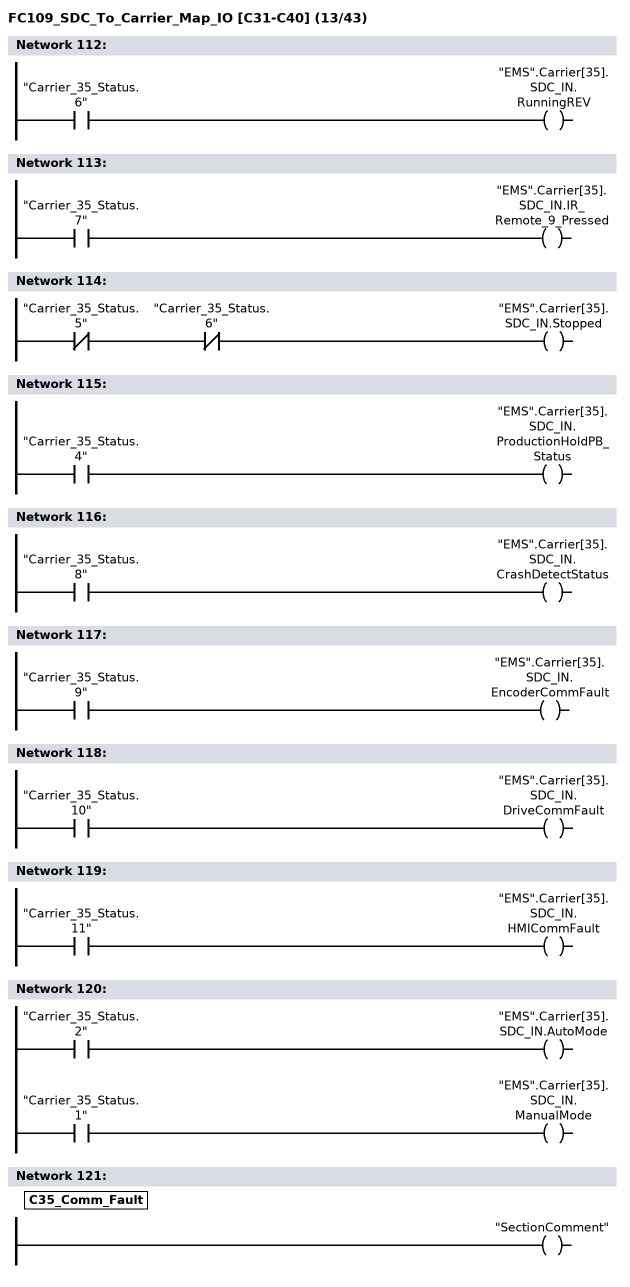
   RUNG wire#powerrail
      Contact( "Carrier_35_Status.6" )
      Coil( "EMS".Carrier[35].SDC_IN.RunningREV )
   END_RUNG
   // the same network as SCL:
   "EMS".Carrier[35].SDC_IN.RunningREV := "Carrier_35_Status.6";
END_REGION

REGION Network 113
   RUNG wire#powerrail
      Contact( "Carrier_35_Status.7" )
      Coil( "EMS".Carrier[35].SDC_IN.IR_Remote_9_Pressed )
   END_RUNG
   // the same network as SCL:
   "EMS".Carrier[35].SDC_IN.IR_Remote_9_Pressed := "Carrier_35_Status.7";
END_REGION

REGION Network 114
   RUNG wire#powerrail
      I_Contact( "Carrier_35_Status.5" )
      I_Contact( "Carrier_35_Status.6" )
      Coil( "EMS".Carrier[35].SDC_IN.Stopped )
   END_RUNG
   // the same network as SCL:
   "EMS".Carrier[35].SDC_IN.Stopped := NOT "Carrier_35_Status.5" AND NOT "Carrier_35_Status.6";
END_REGION

REGION Network 115
   RUNG wire#powerrail
      Contact( "Carrier_35_Status.4" )
      Coil( "EMS".Carrier[35].SDC_IN.ProductionHoldPB_Status )
   END_RUNG
   // the same network as SCL:
   "EMS".Carrier[35].SDC_IN.ProductionHoldPB_Status := "Carrier_35_Status.4";
END_REGION

REGION Network 116
   RUNG wire#powerrail
      Contact( "Carrier_35_Status.8" )
      Coil( "EMS".Carrier[35].SDC_IN.CrashDetectStatus )
   END_RUNG
   // the same network as SCL:
   "EMS".Carrier[35].SDC_IN.CrashDetectStatus := "Carrier_35_Status.8";
END_REGION

REGION Network 117
   RUNG wire#powerrail
      Contact( "Carrier_35_Status.9" )
      Coil( "EMS".Carrier[35].SDC_IN.EncoderCommFault )
   END_RUNG
   // the same network as SCL:
   "EMS".Carrier[35].SDC_IN.EncoderCommFault := "Carrier_35_Status.9";
END_REGION

REGION Network 118
   RUNG wire#powerrail
      Contact( "Carrier_35_Status.10" )
      Coil( "EMS".Carrier[35].SDC_IN.DriveCommFault )
   END_RUNG
   // the same network as SCL:
   "EMS".Carrier[35].SDC_IN.DriveCommFault := "Carrier_35_Status.10";
END_REGION

REGION Network 119
   RUNG wire#powerrail
      Contact( "Carrier_35_Status.11" )
      Coil( "EMS".Carrier[35].SDC_IN.HMICommFault )
   END_RUNG
   // the same network as SCL:
   "EMS".Carrier[35].SDC_IN.HMICommFault := "Carrier_35_Status.11";
END_REGION

REGION Network 120
   RUNG wire#powerrail
      Contact( "Carrier_35_Status.2" )
      Coil( "EMS".Carrier[35].SDC_IN.AutoMode )
   END_RUNG
   RUNG wire#powerrail
      Contact( "Carrier_35_Status.1" )
      Coil( "EMS".Carrier[35].SDC_IN.ManualMode )
   END_RUNG
   // the same network as SCL:
   "EMS".Carrier[35].SDC_IN.AutoMode := "Carrier_35_Status.2";
   "EMS".Carrier[35].SDC_IN.ManualMode := "Carrier_35_Status.1";
END_REGION

REGION Network 121
   Label( C35_Comm_Fault )
   RUNG wire#powerrail
      Coil( "SectionComment" )
   END_RUNG
   // the same network as SCL:
   C35_Comm_Fault:
   "SectionComment" := TRUE;
END_REGION

REGION Network 122
   // **********************************************************************************************************************
   // 
   // Carrier 36 I-Device Data Transfer Interlocks from Carrier to SDC
   // 
   // **********************************************************************************************************************
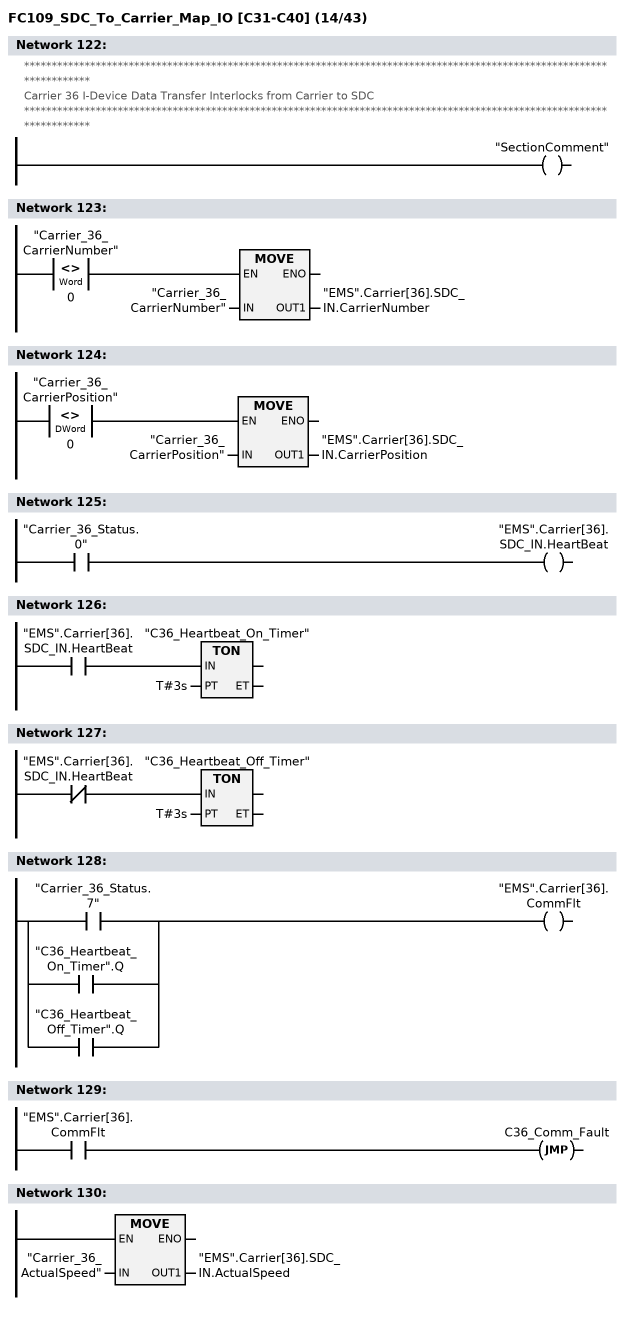
   RUNG wire#powerrail
      Coil( "SectionComment" )
   END_RUNG
   // the same network as SCL:
   "SectionComment" := TRUE;
END_REGION

REGION Network 123
   RUNG wire#powerrail
      { S7_Templates := "SrcType := Word" } NE_Contact(in1 := "Carrier_36_CarrierNumber", in2 := 0)
      Move(in := "Carrier_36_CarrierNumber", out1 => "EMS".Carrier[36].SDC_IN.CarrierNumber)
   END_RUNG
   // the same network as SCL:
   IF "Carrier_36_CarrierNumber" <> 0 THEN
       "EMS".Carrier[36].SDC_IN.CarrierNumber := "Carrier_36_CarrierNumber";
   END_IF;
END_REGION

REGION Network 124
   RUNG wire#powerrail
      { S7_Templates := "SrcType := DWord" } NE_Contact(in1 := "Carrier_36_CarrierPosition", in2 := 0)
      Move(in := "Carrier_36_CarrierPosition", out1 => "EMS".Carrier[36].SDC_IN.CarrierPosition)
   END_RUNG
   // the same network as SCL:
   IF "Carrier_36_CarrierPosition" <> 0 THEN
       "EMS".Carrier[36].SDC_IN.CarrierPosition := "Carrier_36_CarrierPosition";
   END_IF;
END_REGION

REGION Network 125
   RUNG wire#powerrail
      Contact( "Carrier_36_Status.0" )
      Coil( "EMS".Carrier[36].SDC_IN.HeartBeat )
   END_RUNG
   // the same network as SCL:
   "EMS".Carrier[36].SDC_IN.HeartBeat := "Carrier_36_Status.0";
END_REGION

REGION Network 126
   "C36_Heartbeat_On_Timer".TON(IN := "EMS".Carrier[36].SDC_IN.HeartBeat, PT := T#3s);
END_REGION

REGION Network 127
   "C36_Heartbeat_Off_Timer".TON(IN := NOT "EMS".Carrier[36].SDC_IN.HeartBeat, PT := T#3s);
END_REGION

REGION Network 128
   RUNG wire#powerrail
      Contact( "Carrier_36_Status.7" )
      wire#w1
      Coil( "EMS".Carrier[36].CommFlt )
   END_RUNG
   RUNG wire#powerrail
      Contact( "C36_Heartbeat_On_Timer".Q )
   END_RUNG wire#w1
   RUNG wire#powerrail
      Contact( "C36_Heartbeat_Off_Timer".Q )
   END_RUNG wire#w1
   // the same network as SCL:
   "EMS".Carrier[36].CommFlt := "Carrier_36_Status.7" OR "C36_Heartbeat_On_Timer".Q OR "C36_Heartbeat_Off_Timer".Q;
END_REGION

REGION Network 129
   RUNG wire#powerrail
      Contact( "EMS".Carrier[36].CommFlt )
      JumpCoil( C36_Comm_Fault )
   END_RUNG
   // the same network as SCL:
   IF "EMS".Carrier[36].CommFlt THEN GOTO C36_Comm_Fault; END_IF;
END_REGION

REGION Network 130
   RUNG wire#powerrail
      Move(in := "Carrier_36_ActualSpeed", out1 => "EMS".Carrier[36].SDC_IN.ActualSpeed)
   END_RUNG
   // the same network as SCL:
   "EMS".Carrier[36].SDC_IN.ActualSpeed := "Carrier_36_ActualSpeed";
END_REGION

REGION Network 131
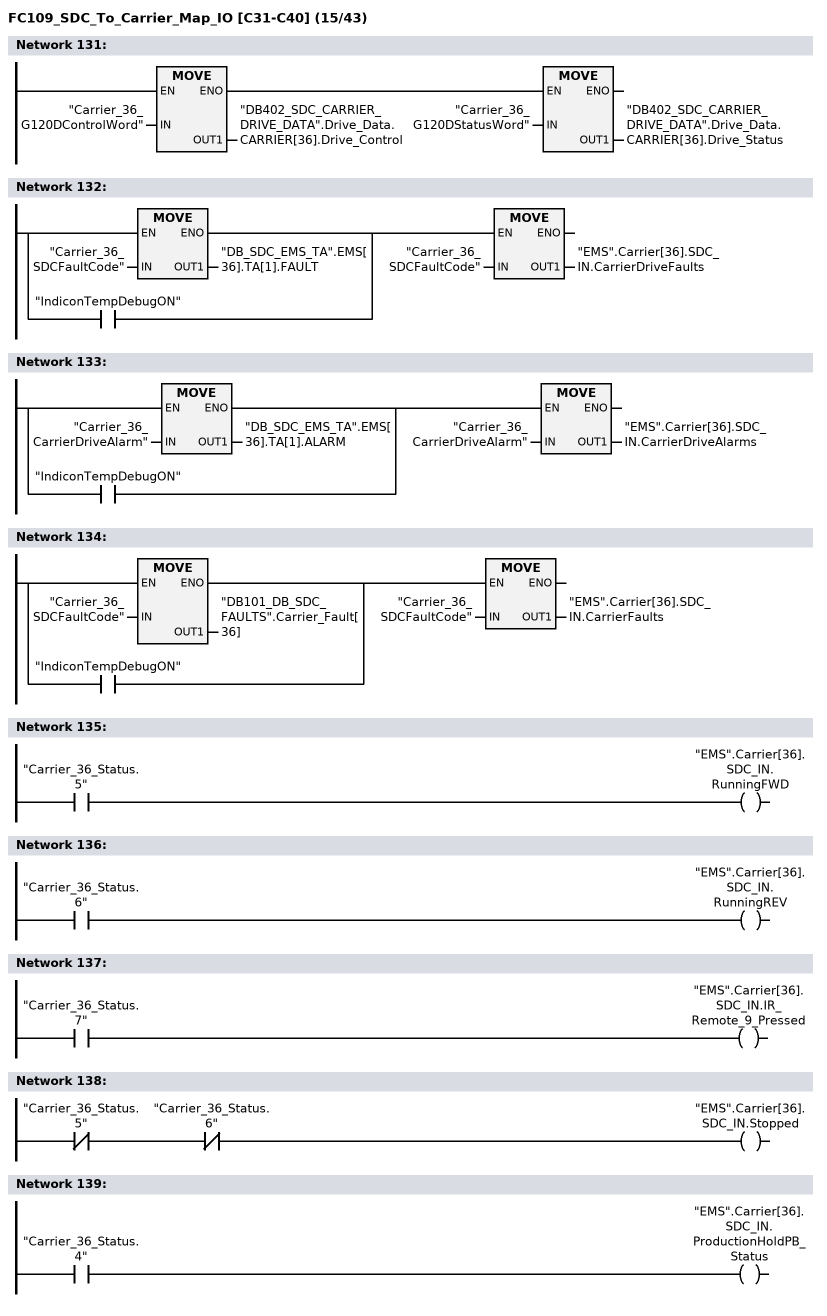
   RUNG wire#powerrail
      Move(in := "Carrier_36_G120DControlWord", out1 => "DB402_SDC_CARRIER_DRIVE_DATA".Drive_Data.CARRIER[36].Drive_Control)
      Move(in := "Carrier_36_G120DStatusWord", out1 => "DB402_SDC_CARRIER_DRIVE_DATA".Drive_Data.CARRIER[36].Drive_Status)
   END_RUNG
   // the same network as SCL:
   "DB402_SDC_CARRIER_DRIVE_DATA".Drive_Data.CARRIER[36].Drive_Control := "Carrier_36_G120DControlWord";
   "DB402_SDC_CARRIER_DRIVE_DATA".Drive_Data.CARRIER[36].Drive_Status := "Carrier_36_G120DStatusWord";
END_REGION

REGION Network 132
   RUNG wire#powerrail
      Move(in := "Carrier_36_SDCFaultCode", out1 => "DB_SDC_EMS_TA".EMS[36].TA[1].FAULT)
      wire#w1
      Move(in := "Carrier_36_SDCFaultCode", out1 => "EMS".Carrier[36].SDC_IN.CarrierDriveFaults)
   END_RUNG
   RUNG wire#powerrail
      Contact( "IndiconTempDebugON" )
   END_RUNG wire#w1
   // the same network as SCL:
   "DB_SDC_EMS_TA".EMS[36].TA[1].FAULT := "Carrier_36_SDCFaultCode";
   IF TRUE OR "IndiconTempDebugON" THEN
       "EMS".Carrier[36].SDC_IN.CarrierDriveFaults := "Carrier_36_SDCFaultCode";
   END_IF;
END_REGION

REGION Network 133
   RUNG wire#powerrail
      Move(in := "Carrier_36_CarrierDriveAlarm", out1 => "DB_SDC_EMS_TA".EMS[36].TA[1].ALARM)
      wire#w1
      Move(in := "Carrier_36_CarrierDriveAlarm", out1 => "EMS".Carrier[36].SDC_IN.CarrierDriveAlarms)
   END_RUNG
   RUNG wire#powerrail
      Contact( "IndiconTempDebugON" )
   END_RUNG wire#w1
   // the same network as SCL:
   "DB_SDC_EMS_TA".EMS[36].TA[1].ALARM := "Carrier_36_CarrierDriveAlarm";
   IF TRUE OR "IndiconTempDebugON" THEN
       "EMS".Carrier[36].SDC_IN.CarrierDriveAlarms := "Carrier_36_CarrierDriveAlarm";
   END_IF;
END_REGION

REGION Network 134
   RUNG wire#powerrail
      Move(in := "Carrier_36_SDCFaultCode", out1 => "DB101_DB_SDC_FAULTS".Carrier_Fault[36])
      wire#w1
      Move(in := "Carrier_36_SDCFaultCode", out1 => "EMS".Carrier[36].SDC_IN.CarrierFaults)
   END_RUNG
   RUNG wire#powerrail
      Contact( "IndiconTempDebugON" )
   END_RUNG wire#w1
   // the same network as SCL:
   "DB101_DB_SDC_FAULTS".Carrier_Fault[36] := "Carrier_36_SDCFaultCode";
   IF TRUE OR "IndiconTempDebugON" THEN
       "EMS".Carrier[36].SDC_IN.CarrierFaults := "Carrier_36_SDCFaultCode";
   END_IF;
END_REGION

REGION Network 135
   RUNG wire#powerrail
      Contact( "Carrier_36_Status.5" )
      Coil( "EMS".Carrier[36].SDC_IN.RunningFWD )
   END_RUNG
   // the same network as SCL:
   "EMS".Carrier[36].SDC_IN.RunningFWD := "Carrier_36_Status.5";
END_REGION

REGION Network 136
   RUNG wire#powerrail
      Contact( "Carrier_36_Status.6" )
      Coil( "EMS".Carrier[36].SDC_IN.RunningREV )
   END_RUNG
   // the same network as SCL:
   "EMS".Carrier[36].SDC_IN.RunningREV := "Carrier_36_Status.6";
END_REGION

REGION Network 137
   RUNG wire#powerrail
      Contact( "Carrier_36_Status.7" )
      Coil( "EMS".Carrier[36].SDC_IN.IR_Remote_9_Pressed )
   END_RUNG
   // the same network as SCL:
   "EMS".Carrier[36].SDC_IN.IR_Remote_9_Pressed := "Carrier_36_Status.7";
END_REGION

REGION Network 138
   RUNG wire#powerrail
      I_Contact( "Carrier_36_Status.5" )
      I_Contact( "Carrier_36_Status.6" )
      Coil( "EMS".Carrier[36].SDC_IN.Stopped )
   END_RUNG
   // the same network as SCL:
   "EMS".Carrier[36].SDC_IN.Stopped := NOT "Carrier_36_Status.5" AND NOT "Carrier_36_Status.6";
END_REGION

REGION Network 139
   RUNG wire#powerrail
      Contact( "Carrier_36_Status.4" )
      Coil( "EMS".Carrier[36].SDC_IN.ProductionHoldPB_Status )
   END_RUNG
   // the same network as SCL:
   "EMS".Carrier[36].SDC_IN.ProductionHoldPB_Status := "Carrier_36_Status.4";
END_REGION

REGION Network 140
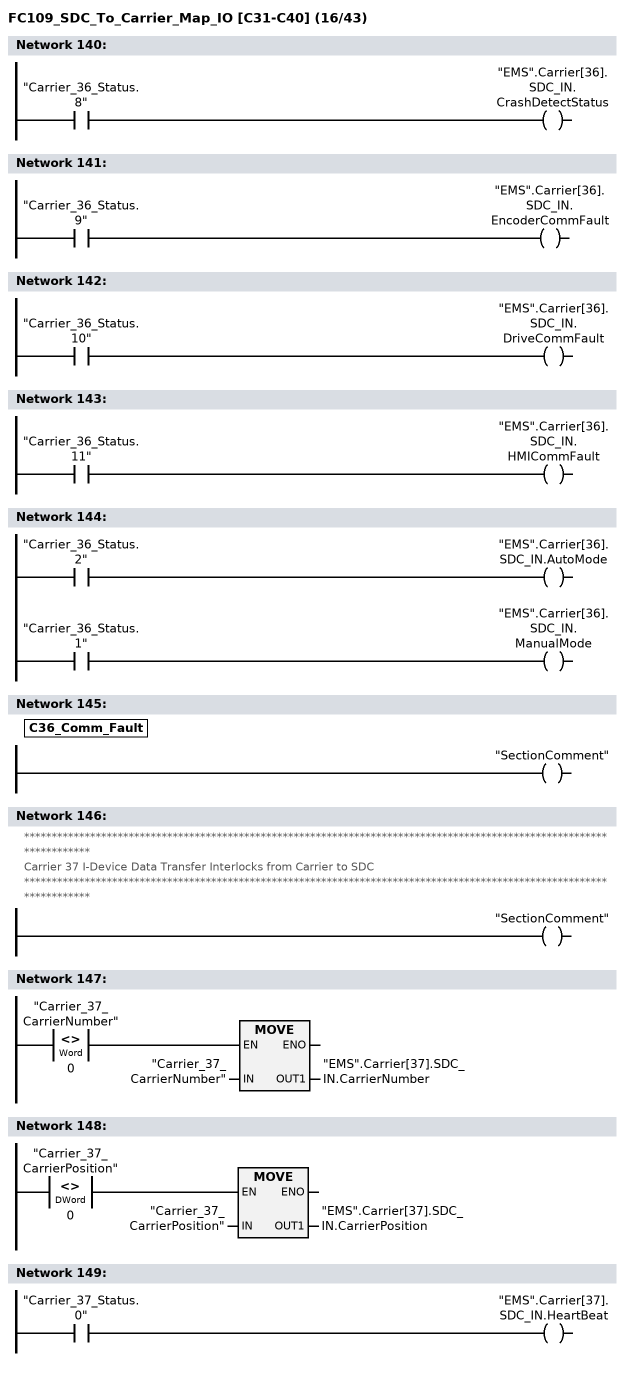
   RUNG wire#powerrail
      Contact( "Carrier_36_Status.8" )
      Coil( "EMS".Carrier[36].SDC_IN.CrashDetectStatus )
   END_RUNG
   // the same network as SCL:
   "EMS".Carrier[36].SDC_IN.CrashDetectStatus := "Carrier_36_Status.8";
END_REGION

REGION Network 141
   RUNG wire#powerrail
      Contact( "Carrier_36_Status.9" )
      Coil( "EMS".Carrier[36].SDC_IN.EncoderCommFault )
   END_RUNG
   // the same network as SCL:
   "EMS".Carrier[36].SDC_IN.EncoderCommFault := "Carrier_36_Status.9";
END_REGION

REGION Network 142
   RUNG wire#powerrail
      Contact( "Carrier_36_Status.10" )
      Coil( "EMS".Carrier[36].SDC_IN.DriveCommFault )
   END_RUNG
   // the same network as SCL:
   "EMS".Carrier[36].SDC_IN.DriveCommFault := "Carrier_36_Status.10";
END_REGION

REGION Network 143
   RUNG wire#powerrail
      Contact( "Carrier_36_Status.11" )
      Coil( "EMS".Carrier[36].SDC_IN.HMICommFault )
   END_RUNG
   // the same network as SCL:
   "EMS".Carrier[36].SDC_IN.HMICommFault := "Carrier_36_Status.11";
END_REGION

REGION Network 144
   RUNG wire#powerrail
      Contact( "Carrier_36_Status.2" )
      Coil( "EMS".Carrier[36].SDC_IN.AutoMode )
   END_RUNG
   RUNG wire#powerrail
      Contact( "Carrier_36_Status.1" )
      Coil( "EMS".Carrier[36].SDC_IN.ManualMode )
   END_RUNG
   // the same network as SCL:
   "EMS".Carrier[36].SDC_IN.AutoMode := "Carrier_36_Status.2";
   "EMS".Carrier[36].SDC_IN.ManualMode := "Carrier_36_Status.1";
END_REGION

REGION Network 145
   Label( C36_Comm_Fault )
   RUNG wire#powerrail
      Coil( "SectionComment" )
   END_RUNG
   // the same network as SCL:
   C36_Comm_Fault:
   "SectionComment" := TRUE;
END_REGION

REGION Network 146
   // **********************************************************************************************************************
   // 
   // Carrier 37 I-Device Data Transfer Interlocks from Carrier to SDC
   // 
   // **********************************************************************************************************************
   RUNG wire#powerrail
      Coil( "SectionComment" )
   END_RUNG
   // the same network as SCL:
   "SectionComment" := TRUE;
END_REGION

REGION Network 147
   RUNG wire#powerrail
      { S7_Templates := "SrcType := Word" } NE_Contact(in1 := "Carrier_37_CarrierNumber", in2 := 0)
      Move(in := "Carrier_37_CarrierNumber", out1 => "EMS".Carrier[37].SDC_IN.CarrierNumber)
   END_RUNG
   // the same network as SCL:
   IF "Carrier_37_CarrierNumber" <> 0 THEN
       "EMS".Carrier[37].SDC_IN.CarrierNumber := "Carrier_37_CarrierNumber";
   END_IF;
END_REGION

REGION Network 148
   RUNG wire#powerrail
      { S7_Templates := "SrcType := DWord" } NE_Contact(in1 := "Carrier_37_CarrierPosition", in2 := 0)
      Move(in := "Carrier_37_CarrierPosition", out1 => "EMS".Carrier[37].SDC_IN.CarrierPosition)
   END_RUNG
   // the same network as SCL:
   IF "Carrier_37_CarrierPosition" <> 0 THEN
       "EMS".Carrier[37].SDC_IN.CarrierPosition := "Carrier_37_CarrierPosition";
   END_IF;
END_REGION

REGION Network 149
   RUNG wire#powerrail
      Contact( "Carrier_37_Status.0" )
      Coil( "EMS".Carrier[37].SDC_IN.HeartBeat )
   END_RUNG
   // the same network as SCL:
   "EMS".Carrier[37].SDC_IN.HeartBeat := "Carrier_37_Status.0";
END_REGION

REGION Network 150
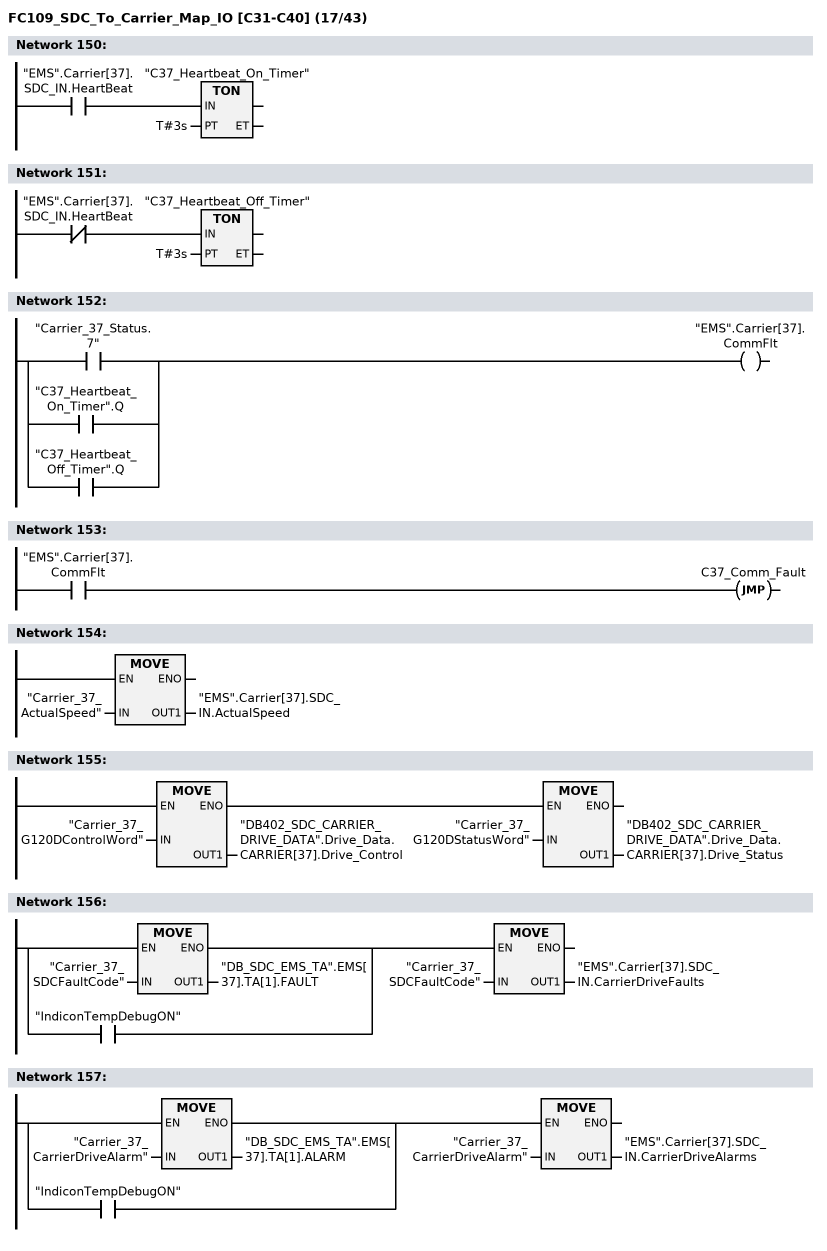
   "C37_Heartbeat_On_Timer".TON(IN := "EMS".Carrier[37].SDC_IN.HeartBeat, PT := T#3s);
END_REGION

REGION Network 151
   "C37_Heartbeat_Off_Timer".TON(IN := NOT "EMS".Carrier[37].SDC_IN.HeartBeat, PT := T#3s);
END_REGION

REGION Network 152
   RUNG wire#powerrail
      Contact( "Carrier_37_Status.7" )
      wire#w1
      Coil( "EMS".Carrier[37].CommFlt )
   END_RUNG
   RUNG wire#powerrail
      Contact( "C37_Heartbeat_On_Timer".Q )
   END_RUNG wire#w1
   RUNG wire#powerrail
      Contact( "C37_Heartbeat_Off_Timer".Q )
   END_RUNG wire#w1
   // the same network as SCL:
   "EMS".Carrier[37].CommFlt := "Carrier_37_Status.7" OR "C37_Heartbeat_On_Timer".Q OR "C37_Heartbeat_Off_Timer".Q;
END_REGION

REGION Network 153
   RUNG wire#powerrail
      Contact( "EMS".Carrier[37].CommFlt )
      JumpCoil( C37_Comm_Fault )
   END_RUNG
   // the same network as SCL:
   IF "EMS".Carrier[37].CommFlt THEN GOTO C37_Comm_Fault; END_IF;
END_REGION

REGION Network 154
   RUNG wire#powerrail
      Move(in := "Carrier_37_ActualSpeed", out1 => "EMS".Carrier[37].SDC_IN.ActualSpeed)
   END_RUNG
   // the same network as SCL:
   "EMS".Carrier[37].SDC_IN.ActualSpeed := "Carrier_37_ActualSpeed";
END_REGION

REGION Network 155
   RUNG wire#powerrail
      Move(in := "Carrier_37_G120DControlWord", out1 => "DB402_SDC_CARRIER_DRIVE_DATA".Drive_Data.CARRIER[37].Drive_Control)
      Move(in := "Carrier_37_G120DStatusWord", out1 => "DB402_SDC_CARRIER_DRIVE_DATA".Drive_Data.CARRIER[37].Drive_Status)
   END_RUNG
   // the same network as SCL:
   "DB402_SDC_CARRIER_DRIVE_DATA".Drive_Data.CARRIER[37].Drive_Control := "Carrier_37_G120DControlWord";
   "DB402_SDC_CARRIER_DRIVE_DATA".Drive_Data.CARRIER[37].Drive_Status := "Carrier_37_G120DStatusWord";
END_REGION

REGION Network 156
   RUNG wire#powerrail
      Move(in := "Carrier_37_SDCFaultCode", out1 => "DB_SDC_EMS_TA".EMS[37].TA[1].FAULT)
      wire#w1
      Move(in := "Carrier_37_SDCFaultCode", out1 => "EMS".Carrier[37].SDC_IN.CarrierDriveFaults)
   END_RUNG
   RUNG wire#powerrail
      Contact( "IndiconTempDebugON" )
   END_RUNG wire#w1
   // the same network as SCL:
   "DB_SDC_EMS_TA".EMS[37].TA[1].FAULT := "Carrier_37_SDCFaultCode";
   IF TRUE OR "IndiconTempDebugON" THEN
       "EMS".Carrier[37].SDC_IN.CarrierDriveFaults := "Carrier_37_SDCFaultCode";
   END_IF;
END_REGION

REGION Network 157
   RUNG wire#powerrail
      Move(in := "Carrier_37_CarrierDriveAlarm", out1 => "DB_SDC_EMS_TA".EMS[37].TA[1].ALARM)
      wire#w1
      Move(in := "Carrier_37_CarrierDriveAlarm", out1 => "EMS".Carrier[37].SDC_IN.CarrierDriveAlarms)
   END_RUNG
   RUNG wire#powerrail
      Contact( "IndiconTempDebugON" )
   END_RUNG wire#w1
   // the same network as SCL:
   "DB_SDC_EMS_TA".EMS[37].TA[1].ALARM := "Carrier_37_CarrierDriveAlarm";
   IF TRUE OR "IndiconTempDebugON" THEN
       "EMS".Carrier[37].SDC_IN.CarrierDriveAlarms := "Carrier_37_CarrierDriveAlarm";
   END_IF;
END_REGION

REGION Network 158
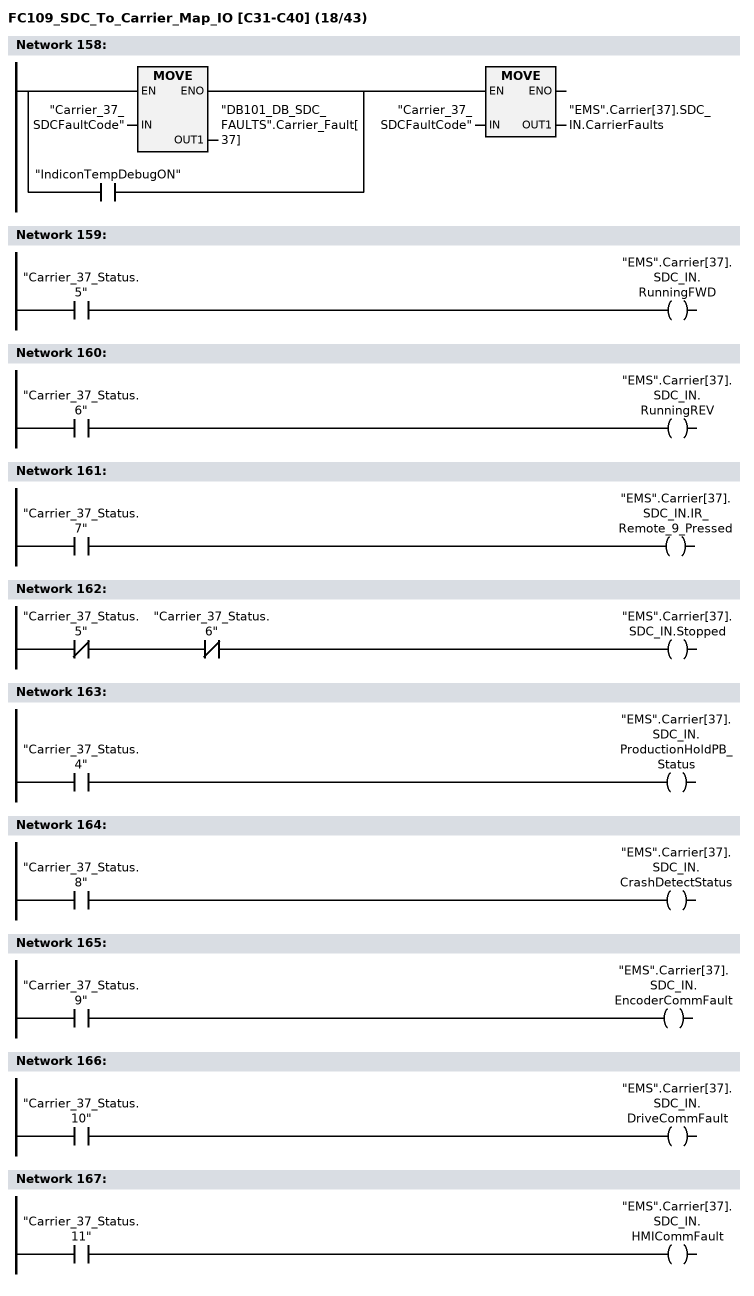
   RUNG wire#powerrail
      Move(in := "Carrier_37_SDCFaultCode", out1 => "DB101_DB_SDC_FAULTS".Carrier_Fault[37])
      wire#w1
      Move(in := "Carrier_37_SDCFaultCode", out1 => "EMS".Carrier[37].SDC_IN.CarrierFaults)
   END_RUNG
   RUNG wire#powerrail
      Contact( "IndiconTempDebugON" )
   END_RUNG wire#w1
   // the same network as SCL:
   "DB101_DB_SDC_FAULTS".Carrier_Fault[37] := "Carrier_37_SDCFaultCode";
   IF TRUE OR "IndiconTempDebugON" THEN
       "EMS".Carrier[37].SDC_IN.CarrierFaults := "Carrier_37_SDCFaultCode";
   END_IF;
END_REGION

REGION Network 159
   RUNG wire#powerrail
      Contact( "Carrier_37_Status.5" )
      Coil( "EMS".Carrier[37].SDC_IN.RunningFWD )
   END_RUNG
   // the same network as SCL:
   "EMS".Carrier[37].SDC_IN.RunningFWD := "Carrier_37_Status.5";
END_REGION

REGION Network 160
   RUNG wire#powerrail
      Contact( "Carrier_37_Status.6" )
      Coil( "EMS".Carrier[37].SDC_IN.RunningREV )
   END_RUNG
   // the same network as SCL:
   "EMS".Carrier[37].SDC_IN.RunningREV := "Carrier_37_Status.6";
END_REGION

REGION Network 161
   RUNG wire#powerrail
      Contact( "Carrier_37_Status.7" )
      Coil( "EMS".Carrier[37].SDC_IN.IR_Remote_9_Pressed )
   END_RUNG
   // the same network as SCL:
   "EMS".Carrier[37].SDC_IN.IR_Remote_9_Pressed := "Carrier_37_Status.7";
END_REGION

REGION Network 162
   RUNG wire#powerrail
      I_Contact( "Carrier_37_Status.5" )
      I_Contact( "Carrier_37_Status.6" )
      Coil( "EMS".Carrier[37].SDC_IN.Stopped )
   END_RUNG
   // the same network as SCL:
   "EMS".Carrier[37].SDC_IN.Stopped := NOT "Carrier_37_Status.5" AND NOT "Carrier_37_Status.6";
END_REGION

REGION Network 163
   RUNG wire#powerrail
      Contact( "Carrier_37_Status.4" )
      Coil( "EMS".Carrier[37].SDC_IN.ProductionHoldPB_Status )
   END_RUNG
   // the same network as SCL:
   "EMS".Carrier[37].SDC_IN.ProductionHoldPB_Status := "Carrier_37_Status.4";
END_REGION

REGION Network 164
   RUNG wire#powerrail
      Contact( "Carrier_37_Status.8" )
      Coil( "EMS".Carrier[37].SDC_IN.CrashDetectStatus )
   END_RUNG
   // the same network as SCL:
   "EMS".Carrier[37].SDC_IN.CrashDetectStatus := "Carrier_37_Status.8";
END_REGION

REGION Network 165
   RUNG wire#powerrail
      Contact( "Carrier_37_Status.9" )
      Coil( "EMS".Carrier[37].SDC_IN.EncoderCommFault )
   END_RUNG
   // the same network as SCL:
   "EMS".Carrier[37].SDC_IN.EncoderCommFault := "Carrier_37_Status.9";
END_REGION

REGION Network 166
   RUNG wire#powerrail
      Contact( "Carrier_37_Status.10" )
      Coil( "EMS".Carrier[37].SDC_IN.DriveCommFault )
   END_RUNG
   // the same network as SCL:
   "EMS".Carrier[37].SDC_IN.DriveCommFault := "Carrier_37_Status.10";
END_REGION

REGION Network 167
   RUNG wire#powerrail
      Contact( "Carrier_37_Status.11" )
      Coil( "EMS".Carrier[37].SDC_IN.HMICommFault )
   END_RUNG
   // the same network as SCL:
   "EMS".Carrier[37].SDC_IN.HMICommFault := "Carrier_37_Status.11";
END_REGION

REGION Network 168
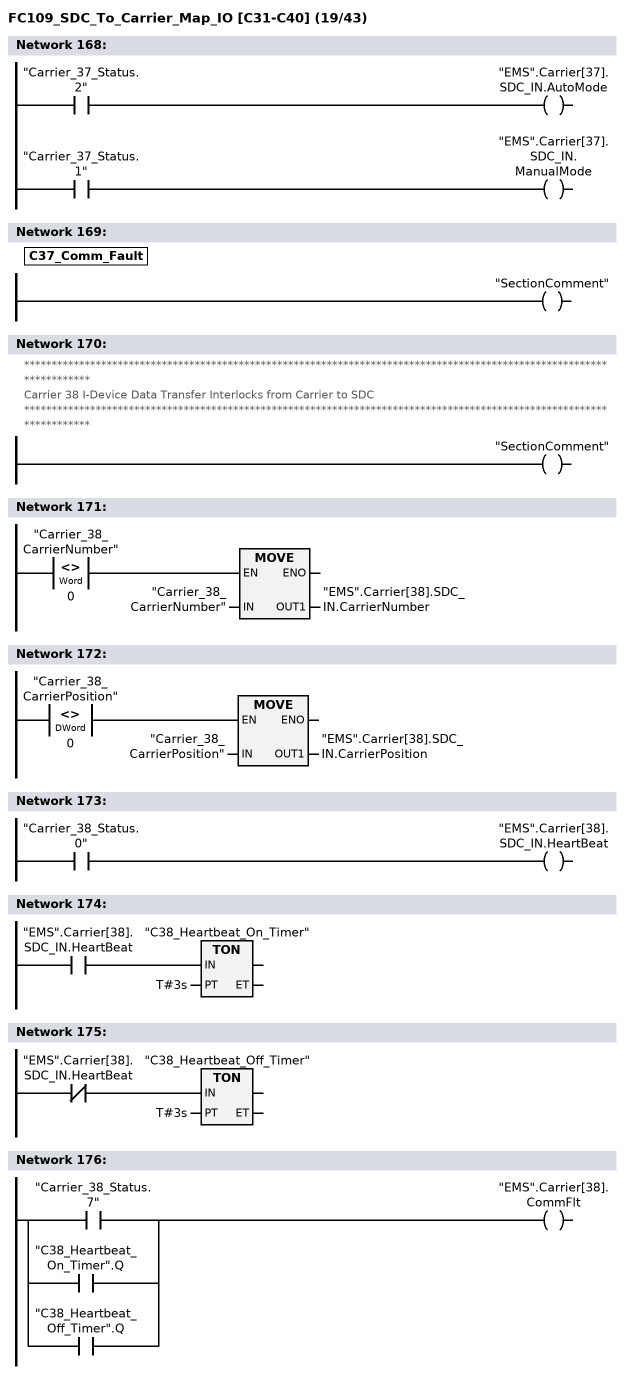
   RUNG wire#powerrail
      Contact( "Carrier_37_Status.2" )
      Coil( "EMS".Carrier[37].SDC_IN.AutoMode )
   END_RUNG
   RUNG wire#powerrail
      Contact( "Carrier_37_Status.1" )
      Coil( "EMS".Carrier[37].SDC_IN.ManualMode )
   END_RUNG
   // the same network as SCL:
   "EMS".Carrier[37].SDC_IN.AutoMode := "Carrier_37_Status.2";
   "EMS".Carrier[37].SDC_IN.ManualMode := "Carrier_37_Status.1";
END_REGION

REGION Network 169
   Label( C37_Comm_Fault )
   RUNG wire#powerrail
      Coil( "SectionComment" )
   END_RUNG
   // the same network as SCL:
   C37_Comm_Fault:
   "SectionComment" := TRUE;
END_REGION

REGION Network 170
   // **********************************************************************************************************************
   // 
   // Carrier 38 I-Device Data Transfer Interlocks from Carrier to SDC
   // 
   // **********************************************************************************************************************
   RUNG wire#powerrail
      Coil( "SectionComment" )
   END_RUNG
   // the same network as SCL:
   "SectionComment" := TRUE;
END_REGION

REGION Network 171
   RUNG wire#powerrail
      { S7_Templates := "SrcType := Word" } NE_Contact(in1 := "Carrier_38_CarrierNumber", in2 := 0)
      Move(in := "Carrier_38_CarrierNumber", out1 => "EMS".Carrier[38].SDC_IN.CarrierNumber)
   END_RUNG
   // the same network as SCL:
   IF "Carrier_38_CarrierNumber" <> 0 THEN
       "EMS".Carrier[38].SDC_IN.CarrierNumber := "Carrier_38_CarrierNumber";
   END_IF;
END_REGION

REGION Network 172
   RUNG wire#powerrail
      { S7_Templates := "SrcType := DWord" } NE_Contact(in1 := "Carrier_38_CarrierPosition", in2 := 0)
      Move(in := "Carrier_38_CarrierPosition", out1 => "EMS".Carrier[38].SDC_IN.CarrierPosition)
   END_RUNG
   // the same network as SCL:
   IF "Carrier_38_CarrierPosition" <> 0 THEN
       "EMS".Carrier[38].SDC_IN.CarrierPosition := "Carrier_38_CarrierPosition";
   END_IF;
END_REGION

REGION Network 173
   RUNG wire#powerrail
      Contact( "Carrier_38_Status.0" )
      Coil( "EMS".Carrier[38].SDC_IN.HeartBeat )
   END_RUNG
   // the same network as SCL:
   "EMS".Carrier[38].SDC_IN.HeartBeat := "Carrier_38_Status.0";
END_REGION

REGION Network 174
   "C38_Heartbeat_On_Timer".TON(IN := "EMS".Carrier[38].SDC_IN.HeartBeat, PT := T#3s);
END_REGION

REGION Network 175
   "C38_Heartbeat_Off_Timer".TON(IN := NOT "EMS".Carrier[38].SDC_IN.HeartBeat, PT := T#3s);
END_REGION

REGION Network 176
   RUNG wire#powerrail
      Contact( "Carrier_38_Status.7" )
      wire#w1
      Coil( "EMS".Carrier[38].CommFlt )
   END_RUNG
   RUNG wire#powerrail
      Contact( "C38_Heartbeat_On_Timer".Q )
   END_RUNG wire#w1
   RUNG wire#powerrail
      Contact( "C38_Heartbeat_Off_Timer".Q )
   END_RUNG wire#w1
   // the same network as SCL:
   "EMS".Carrier[38].CommFlt := "Carrier_38_Status.7" OR "C38_Heartbeat_On_Timer".Q OR "C38_Heartbeat_Off_Timer".Q;
END_REGION

REGION Network 177
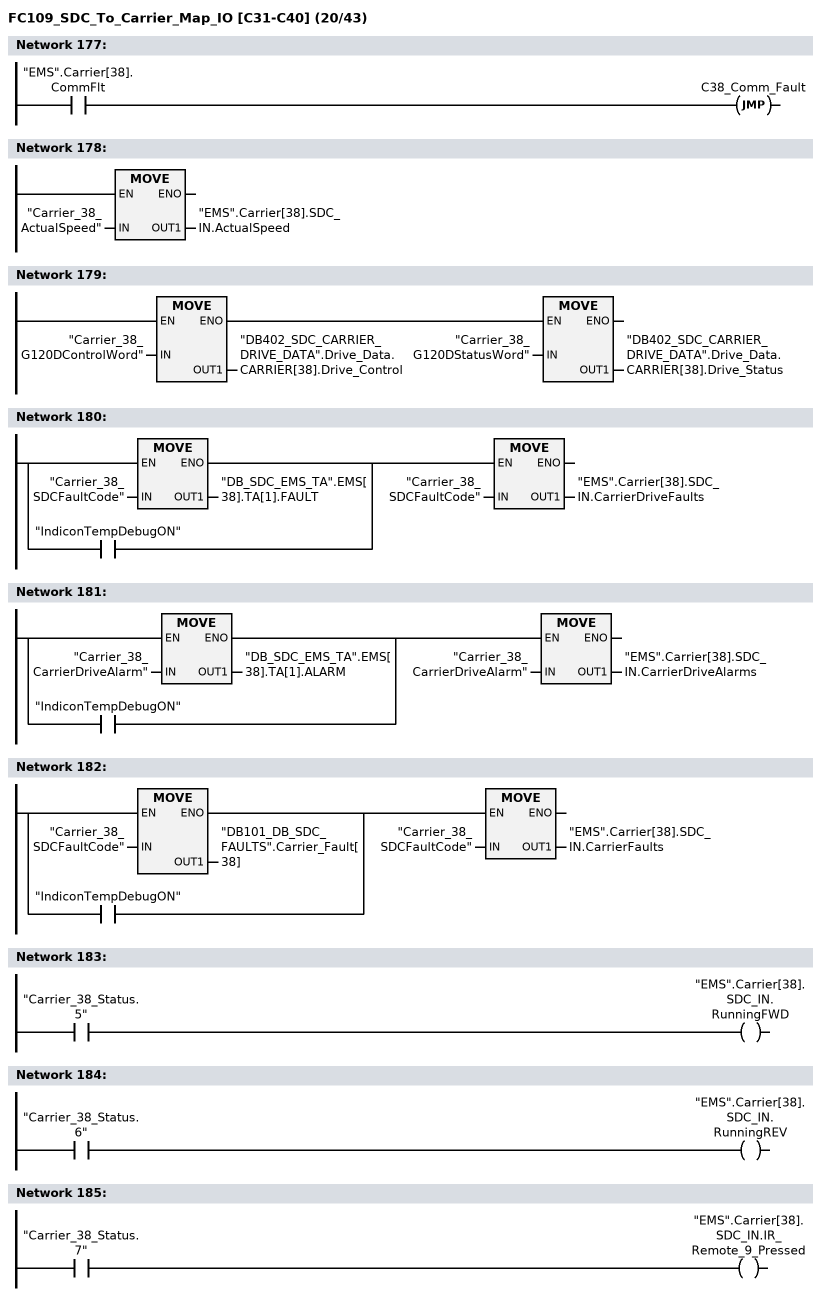
   RUNG wire#powerrail
      Contact( "EMS".Carrier[38].CommFlt )
      JumpCoil( C38_Comm_Fault )
   END_RUNG
   // the same network as SCL:
   IF "EMS".Carrier[38].CommFlt THEN GOTO C38_Comm_Fault; END_IF;
END_REGION

REGION Network 178
   RUNG wire#powerrail
      Move(in := "Carrier_38_ActualSpeed", out1 => "EMS".Carrier[38].SDC_IN.ActualSpeed)
   END_RUNG
   // the same network as SCL:
   "EMS".Carrier[38].SDC_IN.ActualSpeed := "Carrier_38_ActualSpeed";
END_REGION

REGION Network 179
   RUNG wire#powerrail
      Move(in := "Carrier_38_G120DControlWord", out1 => "DB402_SDC_CARRIER_DRIVE_DATA".Drive_Data.CARRIER[38].Drive_Control)
      Move(in := "Carrier_38_G120DStatusWord", out1 => "DB402_SDC_CARRIER_DRIVE_DATA".Drive_Data.CARRIER[38].Drive_Status)
   END_RUNG
   // the same network as SCL:
   "DB402_SDC_CARRIER_DRIVE_DATA".Drive_Data.CARRIER[38].Drive_Control := "Carrier_38_G120DControlWord";
   "DB402_SDC_CARRIER_DRIVE_DATA".Drive_Data.CARRIER[38].Drive_Status := "Carrier_38_G120DStatusWord";
END_REGION

REGION Network 180
   RUNG wire#powerrail
      Move(in := "Carrier_38_SDCFaultCode", out1 => "DB_SDC_EMS_TA".EMS[38].TA[1].FAULT)
      wire#w1
      Move(in := "Carrier_38_SDCFaultCode", out1 => "EMS".Carrier[38].SDC_IN.CarrierDriveFaults)
   END_RUNG
   RUNG wire#powerrail
      Contact( "IndiconTempDebugON" )
   END_RUNG wire#w1
   // the same network as SCL:
   "DB_SDC_EMS_TA".EMS[38].TA[1].FAULT := "Carrier_38_SDCFaultCode";
   IF TRUE OR "IndiconTempDebugON" THEN
       "EMS".Carrier[38].SDC_IN.CarrierDriveFaults := "Carrier_38_SDCFaultCode";
   END_IF;
END_REGION
